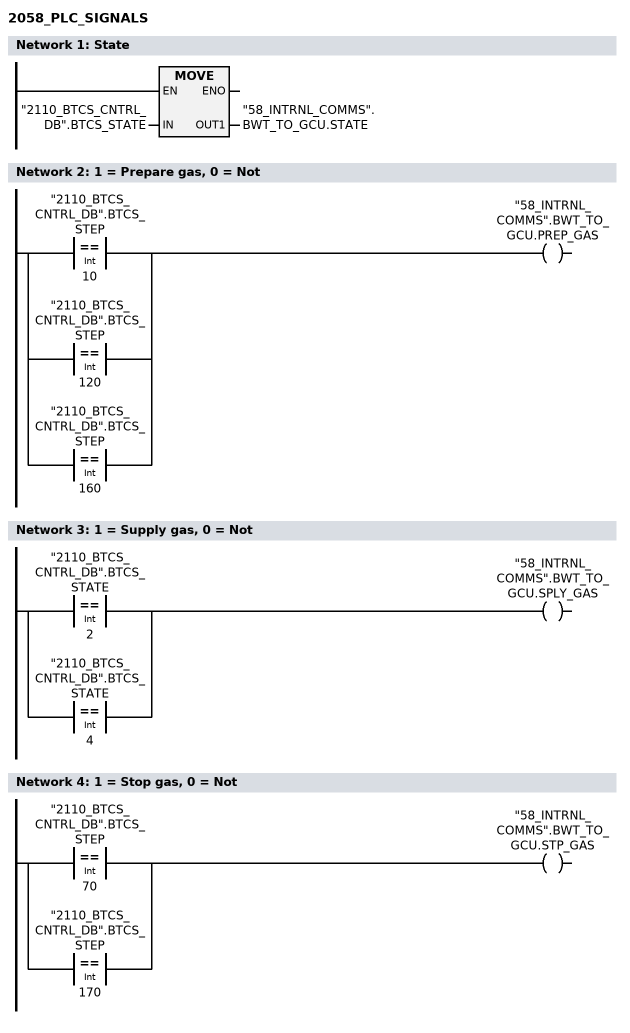
   RUNG wire#powerrail
      Move(in := "2110_BTCS_CNTRL_DB".BTCS_STATE, out1 => "58_INTRNL_COMMS".BWT_TO_GCU.STATE)
   END_RUNG
   // the same network as SCL:
   "58_INTRNL_COMMS".BWT_TO_GCU.STATE := "2110_BTCS_CNTRL_DB".BTCS_STATE;
END_REGION

REGION Network 2: 1 = Prepare gas, 0 = Not
   RUNG wire#powerrail
      { S7_Templates := "SrcType := Int" } EQ_Contact(in1 := "2110_BTCS_CNTRL_DB".BTCS_STEP, in2 := 10)
      wire#w1
      Coil( "58_INTRNL_COMMS".BWT_TO_GCU.PREP_GAS )
   END_RUNG
   RUNG wire#powerrail
      { S7_Templates := "SrcType := Int" } EQ_Contact(in1 := "2110_BTCS_CNTRL_DB".BTCS_STEP, in2 := 120)
   END_RUNG wire#w1
   RUNG wire#powerrail
      { S7_Templates := "SrcType := Int" } EQ_Contact(in1 := "2110_BTCS_CNTRL_DB".BTCS_STEP, in2 := 160)
   END_RUNG wire#w1
   // the same network as SCL:
   "58_INTRNL_COMMS".BWT_TO_GCU.PREP_GAS := ("2110_BTCS_CNTRL_DB".BTCS_STEP = 10) OR ("2110_BTCS_CNTRL_DB".BTCS_STEP = 120) OR ("2110_BTCS_CNTRL_DB".BTCS_STEP = 160);
END_REGION

REGION Network 3: 1 = Supply gas, 0 = Not
   RUNG wire#powerrail
      { S7_Templates := "SrcType := Int" } EQ_Contact(in1 := "2110_BTCS_CNTRL_DB".BTCS_STATE, in2 := 2)
      wire#w1
      Coil( "58_INTRNL_COMMS".BWT_TO_GCU.SPLY_GAS )
   END_RUNG
   RUNG wire#powerrail
      { S7_Templates := "SrcType := Int" } EQ_Contact(in1 := "2110_BTCS_CNTRL_DB".BTCS_STATE, in2 := 4)
   END_RUNG wire#w1
   // the same network as SCL:
   "58_INTRNL_COMMS".BWT_TO_GCU.SPLY_GAS := ("2110_BTCS_CNTRL_DB".BTCS_STATE = 2) OR ("2110_BTCS_CNTRL_DB".BTCS_STATE = 4);
END_REGION

REGION Network 4: 1 = Stop gas, 0 = Not
   RUNG wire#powerrail
      { S7_Templates := "SrcType := Int" } EQ_Contact(in1 := "2110_BTCS_CNTRL_DB".BTCS_STEP, in2 := 70)
      wire#w1
      Coil( "58_INTRNL_COMMS".BWT_TO_GCU.STP_GAS )
   END_RUNG
   RUNG wire#powerrail
      { S7_Templates := "SrcType := Int" } EQ_Contact(in1 := "2110_BTCS_CNTRL_DB".BTCS_STEP, in2 := 170)
   END_RUNG wire#w1
   // the same network as SCL:
   "58_INTRNL_COMMS".BWT_TO_GCU.STP_GAS := ("2110_BTCS_CNTRL_DB".BTCS_STEP = 70) OR ("2110_BTCS_CNTRL_DB".BTCS_STEP = 170);
END_REGION
END_FUNCTION

// folder: 2000 - 2999 BTCS System/2060 - 2069 Alarm & Status Handling

FUNCTION "2060_Alarms" : Void   // FC2060, LAD
TITLE = Alarm Processing
{ S7_Optimized_Access := 'TRUE' }
AUTHOR : JRS
VERSION : 0.1
// To determine alarm conditions
   VAR_TEMP   // added for the SCL form of the ladder/FBD networks
      _w1 : Bool;
   END_VAR
BEGIN

REGION Network 1: DB2060.DBX3.0 = FPT CV422 GTT FPT Fault
   // BTCS_ALARM_WORD_02_BIT_8
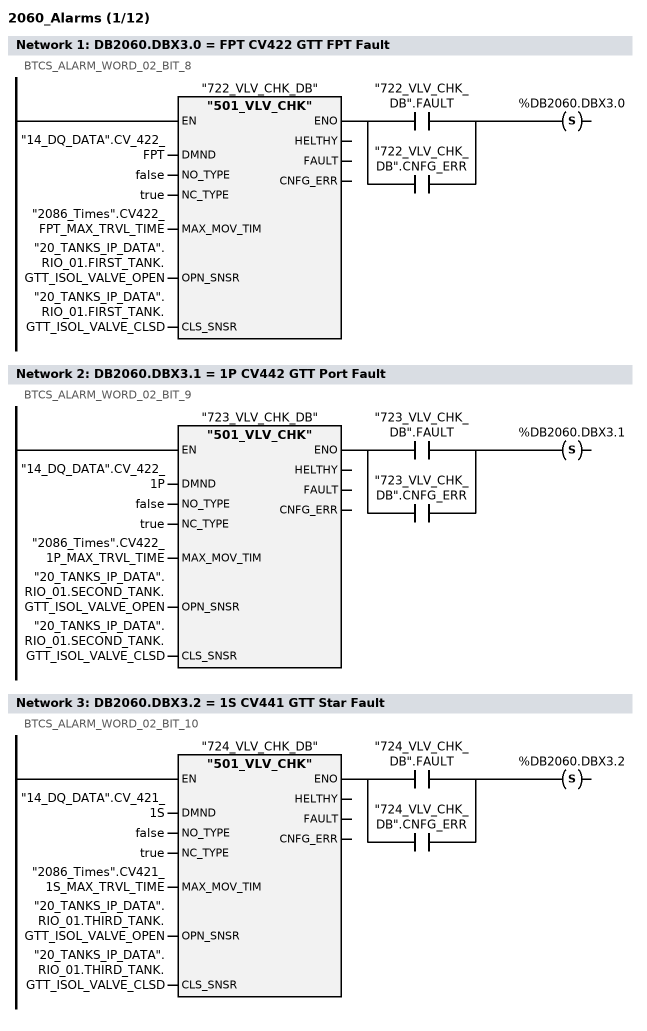
   RUNG wire#powerrail
      "722_VLV_CHK_DB"(DMND := "14_DQ_DATA".CV_422_FPT, NO_TYPE := false, NC_TYPE := true, MAX_MOV_TIM := "2086_Times".CV422_FPT_MAX_TRVL_TIME, OPN_SNSR := "20_TANKS_IP_DATA".RIO_01.FIRST_TANK.GTT_ISOL_VALVE_OPEN, CLS_SNSR := "20_TANKS_IP_DATA".RIO_01.FIRST_TANK.GTT_ISOL_VALVE_CLSD, HELTHY =>, FAULT =>, CNFG_ERR =>)
      wire#w1
      Contact( "722_VLV_CHK_DB".FAULT )
      wire#w2
      S_Coil( %DB2060.DBX3.0 )
   END_RUNG
   RUNG wire#w1
      Contact( "722_VLV_CHK_DB".CNFG_ERR )
   END_RUNG wire#w2
   // the same network as SCL:
   "722_VLV_CHK_DB"(DMND := "14_DQ_DATA".CV_422_FPT,   // "501_VLV_CHK"
                    NO_TYPE := false,
                    NC_TYPE := true,
                    MAX_MOV_TIM := "2086_Times".CV422_FPT_MAX_TRVL_TIME,
                    OPN_SNSR := "20_TANKS_IP_DATA".RIO_01.FIRST_TANK.GTT_ISOL_VALVE_OPEN,
                    CLS_SNSR := "20_TANKS_IP_DATA".RIO_01.FIRST_TANK.GTT_ISOL_VALVE_CLSD,
                    ENO => #_w1);
   IF #_w1 AND ("722_VLV_CHK_DB".FAULT OR "722_VLV_CHK_DB".CNFG_ERR) THEN %DB2060.DBX3.0 := TRUE; END_IF;
END_REGION

REGION Network 2: DB2060.DBX3.1 = 1P CV442 GTT Port Fault
   // BTCS_ALARM_WORD_02_BIT_9
   RUNG wire#powerrail
      "723_VLV_CHK_DB"(DMND := "14_DQ_DATA".CV_422_1P, NO_TYPE := false, NC_TYPE := true, MAX_MOV_TIM := "2086_Times".CV422_1P_MAX_TRVL_TIME, OPN_SNSR := "20_TANKS_IP_DATA".RIO_01.SECOND_TANK.GTT_ISOL_VALVE_OPEN, CLS_SNSR := "20_TANKS_IP_DATA".RIO_01.SECOND_TANK.GTT_ISOL_VALVE_CLSD, HELTHY =>, FAULT =>, CNFG_ERR =>)
      wire#w1
      Contact( "723_VLV_CHK_DB".FAULT )
      wire#w2
      S_Coil( %DB2060.DBX3.1 )
   END_RUNG
   RUNG wire#w1
      Contact( "723_VLV_CHK_DB".CNFG_ERR )
   END_RUNG wire#w2
   // the same network as SCL:
   "723_VLV_CHK_DB"(DMND := "14_DQ_DATA".CV_422_1P,   // "501_VLV_CHK"
                    NO_TYPE := false,
                    NC_TYPE := true,
                    MAX_MOV_TIM := "2086_Times".CV422_1P_MAX_TRVL_TIME,
                    OPN_SNSR := "20_TANKS_IP_DATA".RIO_01.SECOND_TANK.GTT_ISOL_VALVE_OPEN,
                    CLS_SNSR := "20_TANKS_IP_DATA".RIO_01.SECOND_TANK.GTT_ISOL_VALVE_CLSD,
                    ENO => #_w1);
   IF #_w1 AND ("723_VLV_CHK_DB".FAULT OR "723_VLV_CHK_DB".CNFG_ERR) THEN %DB2060.DBX3.1 := TRUE; END_IF;
END_REGION

REGION Network 3: DB2060.DBX3.2 = 1S CV441 GTT Star Fault
   // BTCS_ALARM_WORD_02_BIT_10
   RUNG wire#powerrail
      "724_VLV_CHK_DB"(DMND := "14_DQ_DATA".CV_421_1S, NO_TYPE := false, NC_TYPE := true, MAX_MOV_TIM := "2086_Times".CV421_1S_MAX_TRVL_TIME, OPN_SNSR := "20_TANKS_IP_DATA".RIO_01.THIRD_TANK.GTT_ISOL_VALVE_OPEN, CLS_SNSR := "20_TANKS_IP_DATA".RIO_01.THIRD_TANK.GTT_ISOL_VALVE_CLSD, HELTHY =>, FAULT =>, CNFG_ERR =>)
      wire#w1
      Contact( "724_VLV_CHK_DB".FAULT )
      wire#w2
      S_Coil( %DB2060.DBX3.2 )
   END_RUNG
   RUNG wire#w1
      Contact( "724_VLV_CHK_DB".CNFG_ERR )
   END_RUNG wire#w2
   // the same network as SCL:
   "724_VLV_CHK_DB"(DMND := "14_DQ_DATA".CV_421_1S,   // "501_VLV_CHK"
                    NO_TYPE := false,
                    NC_TYPE := true,
                    MAX_MOV_TIM := "2086_Times".CV421_1S_MAX_TRVL_TIME,
                    OPN_SNSR := "20_TANKS_IP_DATA".RIO_01.THIRD_TANK.GTT_ISOL_VALVE_OPEN,
                    CLS_SNSR := "20_TANKS_IP_DATA".RIO_01.THIRD_TANK.GTT_ISOL_VALVE_CLSD,
                    ENO => #_w1);
   IF #_w1 AND ("724_VLV_CHK_DB".FAULT OR "724_VLV_CHK_DB".CNFG_ERR) THEN %DB2060.DBX3.2 := TRUE; END_IF;
END_REGION

REGION Network 4: DB2060.DBX0.0 = 2P CV442 GTT Port Fault
   // BTCS_ALARM_WORD_01_BIT_0
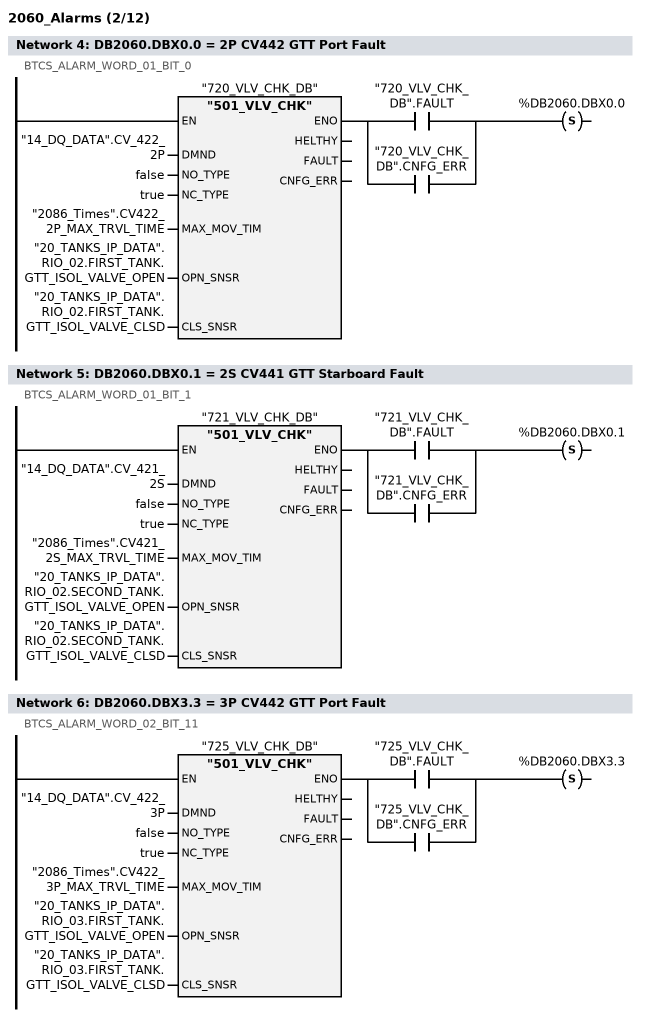
   RUNG wire#powerrail
      "720_VLV_CHK_DB"(DMND := "14_DQ_DATA".CV_422_2P, NO_TYPE := false, NC_TYPE := true, MAX_MOV_TIM := "2086_Times".CV422_2P_MAX_TRVL_TIME, OPN_SNSR := "20_TANKS_IP_DATA".RIO_02.FIRST_TANK.GTT_ISOL_VALVE_OPEN, CLS_SNSR := "20_TANKS_IP_DATA".RIO_02.FIRST_TANK.GTT_ISOL_VALVE_CLSD, HELTHY =>, FAULT =>, CNFG_ERR =>)
      wire#w1
      Contact( "720_VLV_CHK_DB".FAULT )
      wire#w2
      S_Coil( %DB2060.DBX0.0 )
   END_RUNG
   RUNG wire#w1
      Contact( "720_VLV_CHK_DB".CNFG_ERR )
   END_RUNG wire#w2
   // the same network as SCL:
   "720_VLV_CHK_DB"(DMND := "14_DQ_DATA".CV_422_2P,   // "501_VLV_CHK"
                    NO_TYPE := false,
                    NC_TYPE := true,
                    MAX_MOV_TIM := "2086_Times".CV422_2P_MAX_TRVL_TIME,
                    OPN_SNSR := "20_TANKS_IP_DATA".RIO_02.FIRST_TANK.GTT_ISOL_VALVE_OPEN,
                    CLS_SNSR := "20_TANKS_IP_DATA".RIO_02.FIRST_TANK.GTT_ISOL_VALVE_CLSD,
                    ENO => #_w1);
   IF #_w1 AND ("720_VLV_CHK_DB".FAULT OR "720_VLV_CHK_DB".CNFG_ERR) THEN %DB2060.DBX0.0 := TRUE; END_IF;
END_REGION

REGION Network 5: DB2060.DBX0.1 = 2S CV441 GTT Starboard Fault
   // BTCS_ALARM_WORD_01_BIT_1
   RUNG wire#powerrail
      "721_VLV_CHK_DB"(DMND := "14_DQ_DATA".CV_421_2S, NO_TYPE := false, NC_TYPE := true, MAX_MOV_TIM := "2086_Times".CV421_2S_MAX_TRVL_TIME, OPN_SNSR := "20_TANKS_IP_DATA".RIO_02.SECOND_TANK.GTT_ISOL_VALVE_OPEN, CLS_SNSR := "20_TANKS_IP_DATA".RIO_02.SECOND_TANK.GTT_ISOL_VALVE_CLSD, HELTHY =>, FAULT =>, CNFG_ERR =>)
      wire#w1
      Contact( "721_VLV_CHK_DB".FAULT )
      wire#w2
      S_Coil( %DB2060.DBX0.1 )
   END_RUNG
   RUNG wire#w1
      Contact( "721_VLV_CHK_DB".CNFG_ERR )
   END_RUNG wire#w2
   // the same network as SCL:
   "721_VLV_CHK_DB"(DMND := "14_DQ_DATA".CV_421_2S,   // "501_VLV_CHK"
                    NO_TYPE := false,
                    NC_TYPE := true,
                    MAX_MOV_TIM := "2086_Times".CV421_2S_MAX_TRVL_TIME,
                    OPN_SNSR := "20_TANKS_IP_DATA".RIO_02.SECOND_TANK.GTT_ISOL_VALVE_OPEN,
                    CLS_SNSR := "20_TANKS_IP_DATA".RIO_02.SECOND_TANK.GTT_ISOL_VALVE_CLSD,
                    ENO => #_w1);
   IF #_w1 AND ("721_VLV_CHK_DB".FAULT OR "721_VLV_CHK_DB".CNFG_ERR) THEN %DB2060.DBX0.1 := TRUE; END_IF;
END_REGION

REGION Network 6: DB2060.DBX3.3 = 3P CV442 GTT Port Fault
   // BTCS_ALARM_WORD_02_BIT_11
   RUNG wire#powerrail
      "725_VLV_CHK_DB"(DMND := "14_DQ_DATA".CV_422_3P, NO_TYPE := false, NC_TYPE := true, MAX_MOV_TIM := "2086_Times".CV422_3P_MAX_TRVL_TIME, OPN_SNSR := "20_TANKS_IP_DATA".RIO_03.FIRST_TANK.GTT_ISOL_VALVE_OPEN, CLS_SNSR := "20_TANKS_IP_DATA".RIO_03.FIRST_TANK.GTT_ISOL_VALVE_CLSD, HELTHY =>, FAULT =>, CNFG_ERR =>)
      wire#w1
      Contact( "725_VLV_CHK_DB".FAULT )
      wire#w2
      S_Coil( %DB2060.DBX3.3 )
   END_RUNG
   RUNG wire#w1
      Contact( "725_VLV_CHK_DB".CNFG_ERR )
   END_RUNG wire#w2
   // the same network as SCL:
   "725_VLV_CHK_DB"(DMND := "14_DQ_DATA".CV_422_3P,   // "501_VLV_CHK"
                    NO_TYPE := false,
                    NC_TYPE := true,
                    MAX_MOV_TIM := "2086_Times".CV422_3P_MAX_TRVL_TIME,
                    OPN_SNSR := "20_TANKS_IP_DATA".RIO_03.FIRST_TANK.GTT_ISOL_VALVE_OPEN,
                    CLS_SNSR := "20_TANKS_IP_DATA".RIO_03.FIRST_TANK.GTT_ISOL_VALVE_CLSD,
                    ENO => #_w1);
   IF #_w1 AND ("725_VLV_CHK_DB".FAULT OR "725_VLV_CHK_DB".CNFG_ERR) THEN %DB2060.DBX3.3 := TRUE; END_IF;
END_REGION

REGION Network 7: DB2060.DBX3.4 = 3S CV441 GTT Star Fault
   // BTCS_ALARM_WORD_02_BIT_12
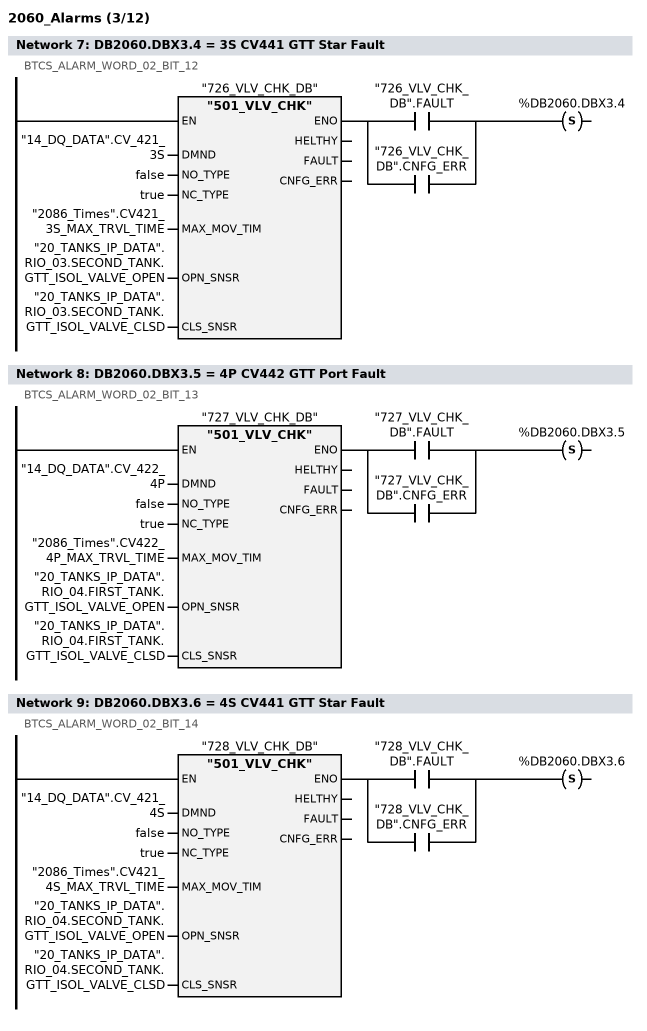
   RUNG wire#powerrail
      "726_VLV_CHK_DB"(DMND := "14_DQ_DATA".CV_421_3S, NO_TYPE := false, NC_TYPE := true, MAX_MOV_TIM := "2086_Times".CV421_3S_MAX_TRVL_TIME, OPN_SNSR := "20_TANKS_IP_DATA".RIO_03.SECOND_TANK.GTT_ISOL_VALVE_OPEN, CLS_SNSR := "20_TANKS_IP_DATA".RIO_03.SECOND_TANK.GTT_ISOL_VALVE_CLSD, HELTHY =>, FAULT =>, CNFG_ERR =>)
      wire#w1
      Contact( "726_VLV_CHK_DB".FAULT )
      wire#w2
      S_Coil( %DB2060.DBX3.4 )
   END_RUNG
   RUNG wire#w1
      Contact( "726_VLV_CHK_DB".CNFG_ERR )
   END_RUNG wire#w2
   // the same network as SCL:
   "726_VLV_CHK_DB"(DMND := "14_DQ_DATA".CV_421_3S,   // "501_VLV_CHK"
                    NO_TYPE := false,
                    NC_TYPE := true,
                    MAX_MOV_TIM := "2086_Times".CV421_3S_MAX_TRVL_TIME,
                    OPN_SNSR := "20_TANKS_IP_DATA".RIO_03.SECOND_TANK.GTT_ISOL_VALVE_OPEN,
                    CLS_SNSR := "20_TANKS_IP_DATA".RIO_03.SECOND_TANK.GTT_ISOL_VALVE_CLSD,
                    ENO => #_w1);
   IF #_w1 AND ("726_VLV_CHK_DB".FAULT OR "726_VLV_CHK_DB".CNFG_ERR) THEN %DB2060.DBX3.4 := TRUE; END_IF;
END_REGION

REGION Network 8: DB2060.DBX3.5 = 4P CV442 GTT Port Fault
   // BTCS_ALARM_WORD_02_BIT_13
   RUNG wire#powerrail
      "727_VLV_CHK_DB"(DMND := "14_DQ_DATA".CV_422_4P, NO_TYPE := false, NC_TYPE := true, MAX_MOV_TIM := "2086_Times".CV422_4P_MAX_TRVL_TIME, OPN_SNSR := "20_TANKS_IP_DATA".RIO_04.FIRST_TANK.GTT_ISOL_VALVE_OPEN, CLS_SNSR := "20_TANKS_IP_DATA".RIO_04.FIRST_TANK.GTT_ISOL_VALVE_CLSD, HELTHY =>, FAULT =>, CNFG_ERR =>)
      wire#w1
      Contact( "727_VLV_CHK_DB".FAULT )
      wire#w2
      S_Coil( %DB2060.DBX3.5 )
   END_RUNG
   RUNG wire#w1
      Contact( "727_VLV_CHK_DB".CNFG_ERR )
   END_RUNG wire#w2
   // the same network as SCL:
   "727_VLV_CHK_DB"(DMND := "14_DQ_DATA".CV_422_4P,   // "501_VLV_CHK"
                    NO_TYPE := false,
                    NC_TYPE := true,
                    MAX_MOV_TIM := "2086_Times".CV422_4P_MAX_TRVL_TIME,
                    OPN_SNSR := "20_TANKS_IP_DATA".RIO_04.FIRST_TANK.GTT_ISOL_VALVE_OPEN,
                    CLS_SNSR := "20_TANKS_IP_DATA".RIO_04.FIRST_TANK.GTT_ISOL_VALVE_CLSD,
                    ENO => #_w1);
   IF #_w1 AND ("727_VLV_CHK_DB".FAULT OR "727_VLV_CHK_DB".CNFG_ERR) THEN %DB2060.DBX3.5 := TRUE; END_IF;
END_REGION

REGION Network 9: DB2060.DBX3.6 = 4S CV441 GTT Star Fault
   // BTCS_ALARM_WORD_02_BIT_14
   RUNG wire#powerrail
      "728_VLV_CHK_DB"(DMND := "14_DQ_DATA".CV_421_4S, NO_TYPE := false, NC_TYPE := true, MAX_MOV_TIM := "2086_Times".CV421_4S_MAX_TRVL_TIME, OPN_SNSR := "20_TANKS_IP_DATA".RIO_04.SECOND_TANK.GTT_ISOL_VALVE_OPEN, CLS_SNSR := "20_TANKS_IP_DATA".RIO_04.SECOND_TANK.GTT_ISOL_VALVE_CLSD, HELTHY =>, FAULT =>, CNFG_ERR =>)
      wire#w1
      Contact( "728_VLV_CHK_DB".FAULT )
      wire#w2
      S_Coil( %DB2060.DBX3.6 )
   END_RUNG
   RUNG wire#w1
      Contact( "728_VLV_CHK_DB".CNFG_ERR )
   END_RUNG wire#w2
   // the same network as SCL:
   "728_VLV_CHK_DB"(DMND := "14_DQ_DATA".CV_421_4S,   // "501_VLV_CHK"
                    NO_TYPE := false,
                    NC_TYPE := true,
                    MAX_MOV_TIM := "2086_Times".CV421_4S_MAX_TRVL_TIME,
                    OPN_SNSR := "20_TANKS_IP_DATA".RIO_04.SECOND_TANK.GTT_ISOL_VALVE_OPEN,
                    CLS_SNSR := "20_TANKS_IP_DATA".RIO_04.SECOND_TANK.GTT_ISOL_VALVE_CLSD,
                    ENO => #_w1);
   IF #_w1 AND ("728_VLV_CHK_DB".FAULT OR "728_VLV_CHK_DB".CNFG_ERR) THEN %DB2060.DBX3.6 := TRUE; END_IF;
END_REGION

REGION Network 10: DB2060.DBX3.7 = 5P CV442 GTT Port Fault
   // BTCS_ALARM_WORD_02_BIT_15
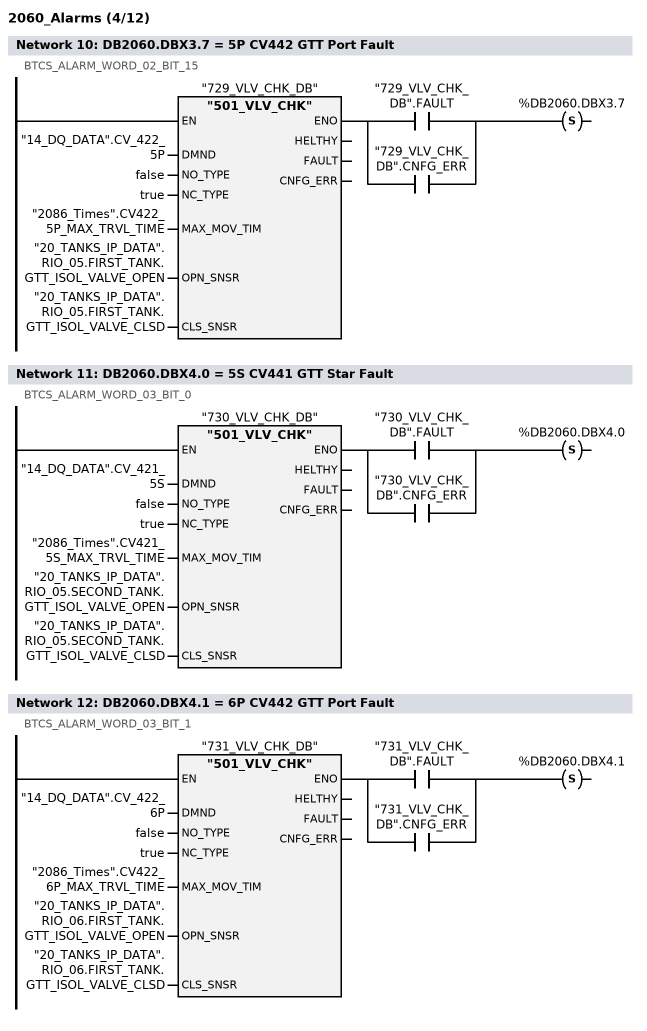
   RUNG wire#powerrail
      "729_VLV_CHK_DB"(DMND := "14_DQ_DATA".CV_422_5P, NO_TYPE := false, NC_TYPE := true, MAX_MOV_TIM := "2086_Times".CV422_5P_MAX_TRVL_TIME, OPN_SNSR := "20_TANKS_IP_DATA".RIO_05.FIRST_TANK.GTT_ISOL_VALVE_OPEN, CLS_SNSR := "20_TANKS_IP_DATA".RIO_05.FIRST_TANK.GTT_ISOL_VALVE_CLSD, HELTHY =>, FAULT =>, CNFG_ERR =>)
      wire#w1
      Contact( "729_VLV_CHK_DB".FAULT )
      wire#w2
      S_Coil( %DB2060.DBX3.7 )
   END_RUNG
   RUNG wire#w1
      Contact( "729_VLV_CHK_DB".CNFG_ERR )
   END_RUNG wire#w2
   // the same network as SCL:
   "729_VLV_CHK_DB"(DMND := "14_DQ_DATA".CV_422_5P,   // "501_VLV_CHK"
                    NO_TYPE := false,
                    NC_TYPE := true,
                    MAX_MOV_TIM := "2086_Times".CV422_5P_MAX_TRVL_TIME,
                    OPN_SNSR := "20_TANKS_IP_DATA".RIO_05.FIRST_TANK.GTT_ISOL_VALVE_OPEN,
                    CLS_SNSR := "20_TANKS_IP_DATA".RIO_05.FIRST_TANK.GTT_ISOL_VALVE_CLSD,
                    ENO => #_w1);
   IF #_w1 AND ("729_VLV_CHK_DB".FAULT OR "729_VLV_CHK_DB".CNFG_ERR) THEN %DB2060.DBX3.7 := TRUE; END_IF;
END_REGION

REGION Network 11: DB2060.DBX4.0 = 5S CV441 GTT Star Fault
   // BTCS_ALARM_WORD_03_BIT_0
   RUNG wire#powerrail
      "730_VLV_CHK_DB"(DMND := "14_DQ_DATA".CV_421_5S, NO_TYPE := false, NC_TYPE := true, MAX_MOV_TIM := "2086_Times".CV421_5S_MAX_TRVL_TIME, OPN_SNSR := "20_TANKS_IP_DATA".RIO_05.SECOND_TANK.GTT_ISOL_VALVE_OPEN, CLS_SNSR := "20_TANKS_IP_DATA".RIO_05.SECOND_TANK.GTT_ISOL_VALVE_CLSD, HELTHY =>, FAULT =>, CNFG_ERR =>)
      wire#w1
      Contact( "730_VLV_CHK_DB".FAULT )
      wire#w2
      S_Coil( %DB2060.DBX4.0 )
   END_RUNG
   RUNG wire#w1
      Contact( "730_VLV_CHK_DB".CNFG_ERR )
   END_RUNG wire#w2
   // the same network as SCL:
   "730_VLV_CHK_DB"(DMND := "14_DQ_DATA".CV_421_5S,   // "501_VLV_CHK"
                    NO_TYPE := false,
                    NC_TYPE := true,
                    MAX_MOV_TIM := "2086_Times".CV421_5S_MAX_TRVL_TIME,
                    OPN_SNSR := "20_TANKS_IP_DATA".RIO_05.SECOND_TANK.GTT_ISOL_VALVE_OPEN,
                    CLS_SNSR := "20_TANKS_IP_DATA".RIO_05.SECOND_TANK.GTT_ISOL_VALVE_CLSD,
                    ENO => #_w1);
   IF #_w1 AND ("730_VLV_CHK_DB".FAULT OR "730_VLV_CHK_DB".CNFG_ERR) THEN %DB2060.DBX4.0 := TRUE; END_IF;
END_REGION

REGION Network 12: DB2060.DBX4.1 = 6P CV442 GTT Port Fault
   // BTCS_ALARM_WORD_03_BIT_1
   RUNG wire#powerrail
      "731_VLV_CHK_DB"(DMND := "14_DQ_DATA".CV_422_6P, NO_TYPE := false, NC_TYPE := true, MAX_MOV_TIM := "2086_Times".CV422_6P_MAX_TRVL_TIME, OPN_SNSR := "20_TANKS_IP_DATA".RIO_06.FIRST_TANK.GTT_ISOL_VALVE_OPEN, CLS_SNSR := "20_TANKS_IP_DATA".RIO_06.FIRST_TANK.GTT_ISOL_VALVE_CLSD, HELTHY =>, FAULT =>, CNFG_ERR =>)
      wire#w1
      Contact( "731_VLV_CHK_DB".FAULT )
      wire#w2
      S_Coil( %DB2060.DBX4.1 )
   END_RUNG
   RUNG wire#w1
      Contact( "731_VLV_CHK_DB".CNFG_ERR )
   END_RUNG wire#w2
   // the same network as SCL:
   "731_VLV_CHK_DB"(DMND := "14_DQ_DATA".CV_422_6P,   // "501_VLV_CHK"
                    NO_TYPE := false,
                    NC_TYPE := true,
                    MAX_MOV_TIM := "2086_Times".CV422_6P_MAX_TRVL_TIME,
                    OPN_SNSR := "20_TANKS_IP_DATA".RIO_06.FIRST_TANK.GTT_ISOL_VALVE_OPEN,
                    CLS_SNSR := "20_TANKS_IP_DATA".RIO_06.FIRST_TANK.GTT_ISOL_VALVE_CLSD,
                    ENO => #_w1);
   IF #_w1 AND ("731_VLV_CHK_DB".FAULT OR "731_VLV_CHK_DB".CNFG_ERR) THEN %DB2060.DBX4.1 := TRUE; END_IF;
END_REGION

REGION Network 13: DB2060.DBX4.2 = 6S CV441 GTT Star Fault
   // BTCS_ALARM_WORD_03_BIT_2
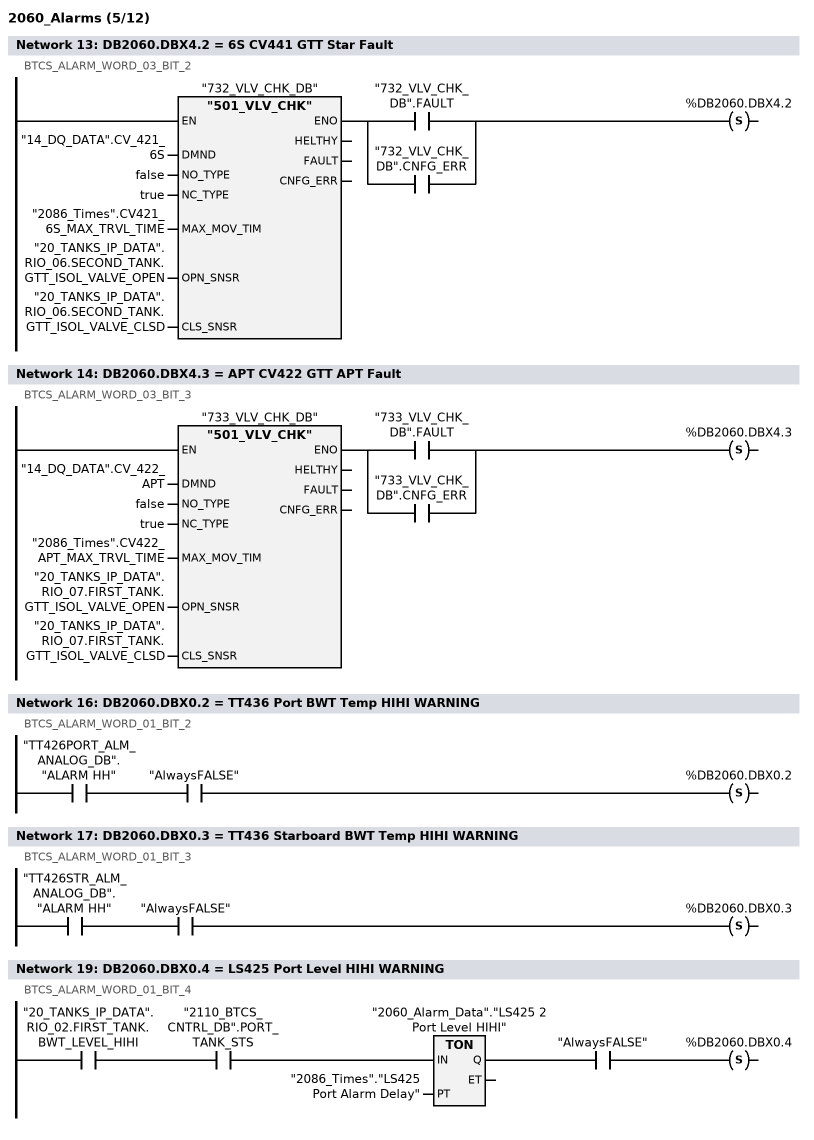
   RUNG wire#powerrail
      "732_VLV_CHK_DB"(DMND := "14_DQ_DATA".CV_421_6S, NO_TYPE := false, NC_TYPE := true, MAX_MOV_TIM := "2086_Times".CV421_6S_MAX_TRVL_TIME, OPN_SNSR := "20_TANKS_IP_DATA".RIO_06.SECOND_TANK.GTT_ISOL_VALVE_OPEN, CLS_SNSR := "20_TANKS_IP_DATA".RIO_06.SECOND_TANK.GTT_ISOL_VALVE_CLSD, HELTHY =>, FAULT =>, CNFG_ERR =>)
      wire#w1
      Contact( "732_VLV_CHK_DB".FAULT )
      wire#w2
      S_Coil( %DB2060.DBX4.2 )
   END_RUNG
   RUNG wire#w1
      Contact( "732_VLV_CHK_DB".CNFG_ERR )
   END_RUNG wire#w2
   // the same network as SCL:
   "732_VLV_CHK_DB"(DMND := "14_DQ_DATA".CV_421_6S,   // "501_VLV_CHK"
                    NO_TYPE := false,
                    NC_TYPE := true,
                    MAX_MOV_TIM := "2086_Times".CV421_6S_MAX_TRVL_TIME,
                    OPN_SNSR := "20_TANKS_IP_DATA".RIO_06.SECOND_TANK.GTT_ISOL_VALVE_OPEN,
                    CLS_SNSR := "20_TANKS_IP_DATA".RIO_06.SECOND_TANK.GTT_ISOL_VALVE_CLSD,
                    ENO => #_w1);
   IF #_w1 AND ("732_VLV_CHK_DB".FAULT OR "732_VLV_CHK_DB".CNFG_ERR) THEN %DB2060.DBX4.2 := TRUE; END_IF;
END_REGION

REGION Network 14: DB2060.DBX4.3 = APT CV422 GTT APT Fault
   // BTCS_ALARM_WORD_03_BIT_3
   RUNG wire#powerrail
      "733_VLV_CHK_DB"(DMND := "14_DQ_DATA".CV_422_APT, NO_TYPE := false, NC_TYPE := true, MAX_MOV_TIM := "2086_Times".CV422_APT_MAX_TRVL_TIME, OPN_SNSR := "20_TANKS_IP_DATA".RIO_07.FIRST_TANK.GTT_ISOL_VALVE_OPEN, CLS_SNSR := "20_TANKS_IP_DATA".RIO_07.FIRST_TANK.GTT_ISOL_VALVE_CLSD, HELTHY =>, FAULT =>, CNFG_ERR =>)
      wire#w1
      Contact( "733_VLV_CHK_DB".FAULT )
      wire#w2
      S_Coil( %DB2060.DBX4.3 )
   END_RUNG
   RUNG wire#w1
      Contact( "733_VLV_CHK_DB".CNFG_ERR )
   END_RUNG wire#w2
   // the same network as SCL:
   "733_VLV_CHK_DB"(DMND := "14_DQ_DATA".CV_422_APT,   // "501_VLV_CHK"
                    NO_TYPE := false,
                    NC_TYPE := true,
                    MAX_MOV_TIM := "2086_Times".CV422_APT_MAX_TRVL_TIME,
                    OPN_SNSR := "20_TANKS_IP_DATA".RIO_07.FIRST_TANK.GTT_ISOL_VALVE_OPEN,
                    CLS_SNSR := "20_TANKS_IP_DATA".RIO_07.FIRST_TANK.GTT_ISOL_VALVE_CLSD,
                    ENO => #_w1);
   IF #_w1 AND ("733_VLV_CHK_DB".FAULT OR "733_VLV_CHK_DB".CNFG_ERR) THEN %DB2060.DBX4.3 := TRUE; END_IF;
END_REGION

REGION Network 16: DB2060.DBX0.2 = TT436 Port BWT Temp HIHI WARNING
   // BTCS_ALARM_WORD_01_BIT_2
   RUNG wire#powerrail
      Contact( "TT426PORT_ALM_ANALOG_DB"."ALARM HH" )
      Contact( "AlwaysFALSE" )
      S_Coil( %DB2060.DBX0.2 )
   END_RUNG
   // the same network as SCL:
   IF "TT426PORT_ALM_ANALOG_DB"."ALARM HH" AND "AlwaysFALSE" THEN %DB2060.DBX0.2 := TRUE; END_IF;
END_REGION

REGION Network 17: DB2060.DBX0.3 = TT436 Starboard BWT Temp HIHI WARNING
   // BTCS_ALARM_WORD_01_BIT_3
   RUNG wire#powerrail
      Contact( "TT426STR_ALM_ANALOG_DB"."ALARM HH" )
      Contact( "AlwaysFALSE" )
      S_Coil( %DB2060.DBX0.3 )
   END_RUNG
   // the same network as SCL:
   IF "TT426STR_ALM_ANALOG_DB"."ALARM HH" AND "AlwaysFALSE" THEN %DB2060.DBX0.3 := TRUE; END_IF;
END_REGION

REGION Network 19: DB2060.DBX0.4 = LS425 Port Level HIHI WARNING
   // BTCS_ALARM_WORD_01_BIT_4
   "2060_Alarm_Data"."LS425 2 Port Level HIHI".TON(IN := "20_TANKS_IP_DATA".RIO_02.FIRST_TANK.BWT_LEVEL_HIHI AND "2110_BTCS_CNTRL_DB".PORT_TANK_STS,
                           PT := "2086_Times"."LS425 Port Alarm Delay");
   IF "2060_Alarm_Data"."LS425 2 Port Level HIHI".Q AND "AlwaysFALSE" THEN %DB2060.DBX0.4 := TRUE; END_IF;
END_REGION

REGION Network 20: DB2060.DBX0.5 = LS425 Starboard Level HIHI WARNING
   // BTCS_ALARM_WORD_01_BIT_5
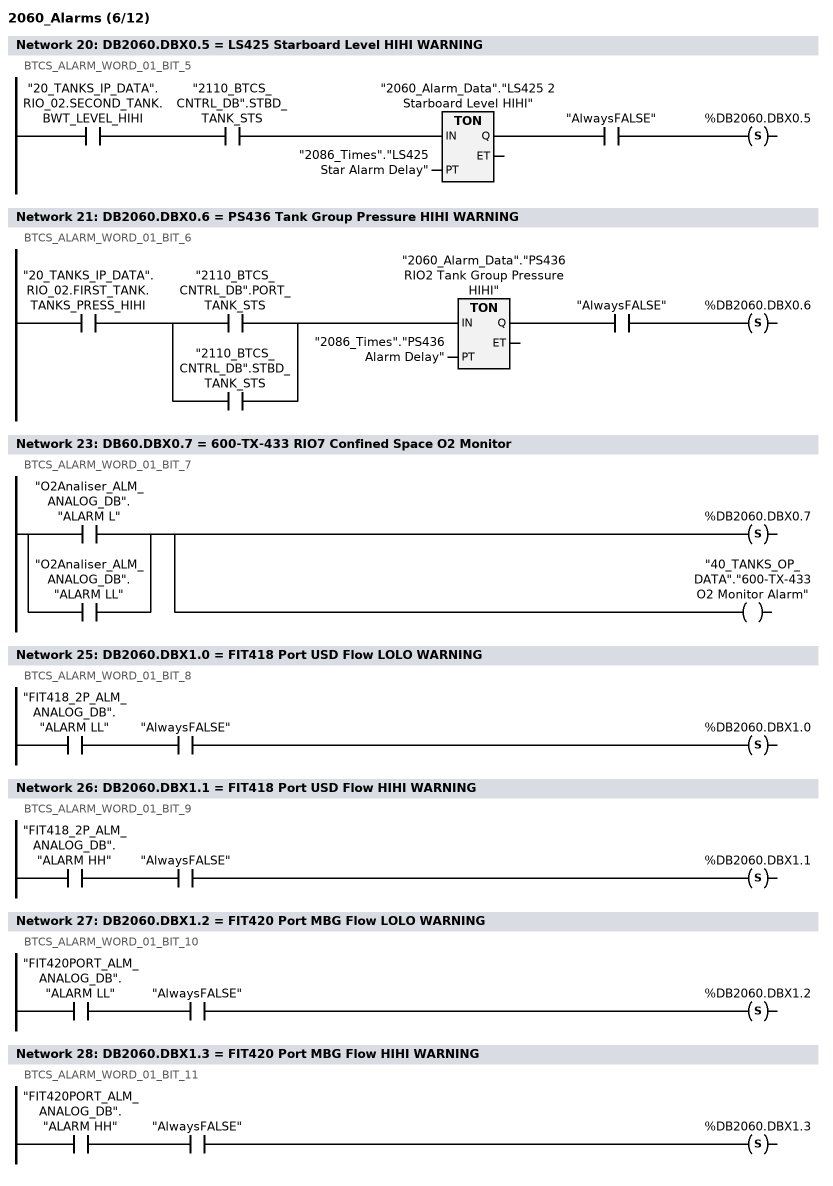
   "2060_Alarm_Data"."LS425 2 Starboard Level HIHI".TON(IN := "20_TANKS_IP_DATA".RIO_02.SECOND_TANK.BWT_LEVEL_HIHI AND "2110_BTCS_CNTRL_DB".STBD_TANK_STS,
                           PT := "2086_Times"."LS425 Star Alarm Delay");
   IF "2060_Alarm_Data"."LS425 2 Starboard Level HIHI".Q AND "AlwaysFALSE" THEN
       %DB2060.DBX0.5 := TRUE;
   END_IF;
END_REGION

REGION Network 21: DB2060.DBX0.6 = PS436 Tank Group Pressure HIHI WARNING
   // BTCS_ALARM_WORD_01_BIT_6
   "2060_Alarm_Data"."PS436 RIO2 Tank Group Pressure HIHI".TON(IN := "20_TANKS_IP_DATA".RIO_02.FIRST_TANK.TANKS_PRESS_HIHI AND ("2110_BTCS_CNTRL_DB".PORT_TANK_STS OR "2110_BTCS_CNTRL_DB".STBD_TANK_STS),
                           PT := "2086_Times"."PS436 Alarm Delay");
   IF "2060_Alarm_Data"."PS436 RIO2 Tank Group Pressure HIHI".Q AND "AlwaysFALSE" THEN
       %DB2060.DBX0.6 := TRUE;
   END_IF;
END_REGION

REGION Network 23: DB60.DBX0.7 = 600-TX-433 RIO7 Confined Space O2 Monitor
   // BTCS_ALARM_WORD_01_BIT_7
   RUNG wire#powerrail
      Contact( "O2Analiser_ALM_ANALOG_DB"."ALARM L" )
      wire#w1
      S_Coil( %DB2060.DBX0.7 )
   END_RUNG
   RUNG wire#powerrail
      Contact( "O2Analiser_ALM_ANALOG_DB"."ALARM LL" )
   END_RUNG wire#w1
   RUNG wire#w1
      Coil( "40_TANKS_OP_DATA"."600-TX-433  O2 Monitor Alarm" )
   END_RUNG
   // the same network as SCL:
   #_w1 := "O2Analiser_ALM_ANALOG_DB"."ALARM L" OR "O2Analiser_ALM_ANALOG_DB"."ALARM LL";
   IF #_w1 THEN %DB2060.DBX0.7 := TRUE; END_IF;
   "40_TANKS_OP_DATA"."600-TX-433  O2 Monitor Alarm" := #_w1;
END_REGION

REGION Network 25: DB2060.DBX1.0 = FIT418 Port USD Flow LOLO WARNING
   // BTCS_ALARM_WORD_01_BIT_8
   RUNG wire#powerrail
      Contact( "FIT418_2P_ALM_ANALOG_DB"."ALARM LL" )
      Contact( "AlwaysFALSE" )
      S_Coil( %DB2060.DBX1.0 )
   END_RUNG
   // the same network as SCL:
   IF "FIT418_2P_ALM_ANALOG_DB"."ALARM LL" AND "AlwaysFALSE" THEN %DB2060.DBX1.0 := TRUE; END_IF;
END_REGION

REGION Network 26: DB2060.DBX1.1 = FIT418 Port USD Flow HIHI WARNING
   // BTCS_ALARM_WORD_01_BIT_9
   RUNG wire#powerrail
      Contact( "FIT418_2P_ALM_ANALOG_DB"."ALARM HH" )
      Contact( "AlwaysFALSE" )
      S_Coil( %DB2060.DBX1.1 )
   END_RUNG
   // the same network as SCL:
   IF "FIT418_2P_ALM_ANALOG_DB"."ALARM HH" AND "AlwaysFALSE" THEN %DB2060.DBX1.1 := TRUE; END_IF;
END_REGION

REGION Network 27: DB2060.DBX1.2 = FIT420 Port MBG Flow LOLO WARNING
   // BTCS_ALARM_WORD_01_BIT_10
   RUNG wire#powerrail
      Contact( "FIT420PORT_ALM_ANALOG_DB"."ALARM LL" )
      Contact( "AlwaysFALSE" )
      S_Coil( %DB2060.DBX1.2 )
   END_RUNG
   // the same network as SCL:
   IF "FIT420PORT_ALM_ANALOG_DB"."ALARM LL" AND "AlwaysFALSE" THEN %DB2060.DBX1.2 := TRUE; END_IF;
END_REGION

REGION Network 28: DB2060.DBX1.3 = FIT420 Port MBG Flow HIHI WARNING
   // BTCS_ALARM_WORD_01_BIT_11
   RUNG wire#powerrail
      Contact( "FIT420PORT_ALM_ANALOG_DB"."ALARM HH" )
      Contact( "AlwaysFALSE" )
      S_Coil( %DB2060.DBX1.3 )
   END_RUNG
   // the same network as SCL:
   IF "FIT420PORT_ALM_ANALOG_DB"."ALARM HH" AND "AlwaysFALSE" THEN %DB2060.DBX1.3 := TRUE; END_IF;
END_REGION

REGION Network 29: DB2060.DBX1.4 = FIT417 Starboard USD Flow LOLO WARNING
   // BTCS_ALARM_WORD_01_BIT_12
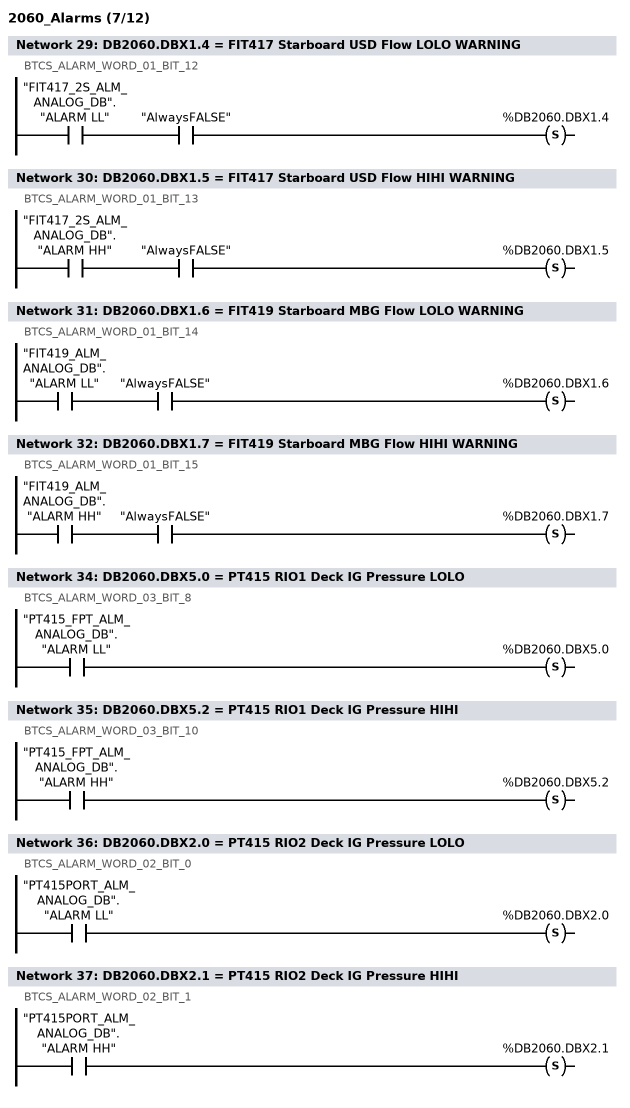
   RUNG wire#powerrail
      Contact( "FIT417_2S_ALM_ANALOG_DB"."ALARM LL" )
      Contact( "AlwaysFALSE" )
      S_Coil( %DB2060.DBX1.4 )
   END_RUNG
   // the same network as SCL:
   IF "FIT417_2S_ALM_ANALOG_DB"."ALARM LL" AND "AlwaysFALSE" THEN %DB2060.DBX1.4 := TRUE; END_IF;
END_REGION

REGION Network 30: DB2060.DBX1.5 = FIT417 Starboard USD Flow HIHI WARNING
   // BTCS_ALARM_WORD_01_BIT_13
   RUNG wire#powerrail
      Contact( "FIT417_2S_ALM_ANALOG_DB"."ALARM HH" )
      Contact( "AlwaysFALSE" )
      S_Coil( %DB2060.DBX1.5 )
   END_RUNG
   // the same network as SCL:
   IF "FIT417_2S_ALM_ANALOG_DB"."ALARM HH" AND "AlwaysFALSE" THEN %DB2060.DBX1.5 := TRUE; END_IF;
END_REGION

REGION Network 31: DB2060.DBX1.6 = FIT419 Starboard MBG Flow LOLO WARNING
   // BTCS_ALARM_WORD_01_BIT_14
   RUNG wire#powerrail
      Contact( "FIT419_ALM_ANALOG_DB"."ALARM LL" )
      Contact( "AlwaysFALSE" )
      S_Coil( %DB2060.DBX1.6 )
   END_RUNG
   // the same network as SCL:
   IF "FIT419_ALM_ANALOG_DB"."ALARM LL" AND "AlwaysFALSE" THEN %DB2060.DBX1.6 := TRUE; END_IF;
END_REGION

REGION Network 32: DB2060.DBX1.7 = FIT419 Starboard MBG Flow HIHI WARNING
   // BTCS_ALARM_WORD_01_BIT_15
   RUNG wire#powerrail
      Contact( "FIT419_ALM_ANALOG_DB"."ALARM HH" )
      Contact( "AlwaysFALSE" )
      S_Coil( %DB2060.DBX1.7 )
   END_RUNG
   // the same network as SCL:
   IF "FIT419_ALM_ANALOG_DB"."ALARM HH" AND "AlwaysFALSE" THEN %DB2060.DBX1.7 := TRUE; END_IF;
END_REGION

REGION Network 34: DB2060.DBX5.0 = PT415 RIO1 Deck IG Pressure LOLO
   // BTCS_ALARM_WORD_03_BIT_8
   RUNG wire#powerrail
      Contact( "PT415_FPT_ALM_ANALOG_DB"."ALARM LL" )
      S_Coil( %DB2060.DBX5.0 )
   END_RUNG
   // the same network as SCL:
   IF "PT415_FPT_ALM_ANALOG_DB"."ALARM LL" THEN %DB2060.DBX5.0 := TRUE; END_IF;
END_REGION

REGION Network 35: DB2060.DBX5.2 = PT415 RIO1 Deck IG Pressure HIHI
   // BTCS_ALARM_WORD_03_BIT_10
   RUNG wire#powerrail
      Contact( "PT415_FPT_ALM_ANALOG_DB"."ALARM HH" )
      S_Coil( %DB2060.DBX5.2 )
   END_RUNG
   // the same network as SCL:
   IF "PT415_FPT_ALM_ANALOG_DB"."ALARM HH" THEN %DB2060.DBX5.2 := TRUE; END_IF;
END_REGION

REGION Network 36: DB2060.DBX2.0 = PT415 RIO2 Deck IG Pressure LOLO
   // BTCS_ALARM_WORD_02_BIT_0
   RUNG wire#powerrail
      Contact( "PT415PORT_ALM_ANALOG_DB"."ALARM LL" )
      S_Coil( %DB2060.DBX2.0 )
   END_RUNG
   // the same network as SCL:
   IF "PT415PORT_ALM_ANALOG_DB"."ALARM LL" THEN %DB2060.DBX2.0 := TRUE; END_IF;
END_REGION

REGION Network 37: DB2060.DBX2.1 = PT415 RIO2 Deck IG Pressure HIHI
   // BTCS_ALARM_WORD_02_BIT_1
   RUNG wire#powerrail
      Contact( "PT415PORT_ALM_ANALOG_DB"."ALARM HH" )
      S_Coil( %DB2060.DBX2.1 )
   END_RUNG
   // the same network as SCL:
   IF "PT415PORT_ALM_ANALOG_DB"."ALARM HH" THEN %DB2060.DBX2.1 := TRUE; END_IF;
END_REGION

REGION Network 38: DB2060.DBX5.3 = PT415 RIO3 Deck IG Pressure LOLO
   // BTCS_ALARM_WORD_03_BIT_11
